// TIA Portal project "Tank_Level_FactoryIO" (V15.1)

(* hardware
DEVICE "S7-1200 station_1"  S7-1200 Station
   slot 0: "Rack_0"  S7-1200 Rack  Rack  V1.0
   slot 1: "PLC_1"  CPU 1214C DC/DC/DC  6ES7 214-1AG40-0XB0  V4.2
DEVICE "HMI_1"  TP1500 Comfort PRO
   slot 0: "HMI_1"  TP1500 Comfort PRO  6AV2 124-0QC24-1AX0  15.1.0.0
   slot 1: "HMI_RT_1"  TP1500 Comfort PRO  6AV2 124-0QC24-1AX0  15.1.0.0
   slot 5: "HMI_1.IE_CP_1"  PROFINET Interface  15.0.1.0
      slot 1: "PROFINET Interface_1"  PROFINET Interface
         slot 1: "Port_1"  Port
         slot 2: "Port_2"  Port
   slot 6: "HMI_1.IE_CP_2"  PROFINET Interface  15.0.1.0
      slot 1: "PROFINET Interface_GBit"  PROFINET Interface
         slot 1: "Port_1"  Port
   slot 7: "HMI_1.MPI/DP_CP_1"  MPI/DP Interface  15.0.1.0
*)

// ===== PLC "PLC_1"  CPU 1214C DC/DC/DC =====

VAR_GLOBAL   // PLC tag table "Default tag table"
   "Raw_Sensor_Sim" AT %MW10 : Int;
   "Level_Normalized" AT %MD20 : Real;
   "Level_CM" AT %MD24 : Real;
   "Fill_Valve" AT %QW30 : Int;
   "Pump_Cmd" AT %Q0.0 : Bool;
   "I_Start" AT %I0.0 : Bool;
   "I_Stop" AT %I0.1 : Bool;
   "System_Active" AT %M0.0 : Bool;
   "Discharge_Valve" AT %Q0.1 : Bool;
   "Sim_Tick" AT %M50.0 : Bool;
   "Level_Input_Raw" AT %IW30 : Int;
   "Discharge_Valve_Analog" AT %QW32 : Int;
   "HMI_Start" AT %M10.0 : Bool;
   "HMI_Stop" AT %M12.0 : Bool;
END_VAR

FUNCTION "Signal Conversion" : Void   // FC1, LAD
{ S7_Optimized_Access := 'TRUE' }
VERSION : 0.1
BEGIN

REGION Network 1: Signal Conversion
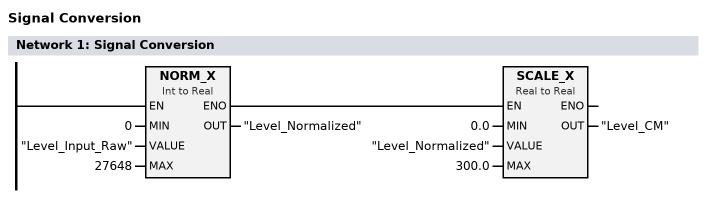
   RUNG wire#powerrail
      { S7_Templates := "[SrcType := Int, DestType := Real]" } Normalize(min := 0, value := "Level_Input_Raw", max := 27648, out => "Level_Normalized")
      { S7_Templates := "[SrcType := Real, DestType := Real]" } Scale(min := 0.0, value := "Level_Normalized", max := 300.0, out => "Level_CM")
   END_RUNG
   // the same network as SCL:
   "Level_Normalized" := NORM_X(MIN := 0, VALUE := "Level_Input_Raw", MAX := 27648);
   "Level_CM" := SCALE_X(MIN := 0.0, VALUE := "Level_Normalized", MAX := 300.0);
END_REGION
END_FUNCTION

FUNCTION "Pump Control" : Void   // FC2, LAD
{ S7_Optimized_Access := 'TRUE' }
VERSION : 0.1
BEGIN

REGION Network 1
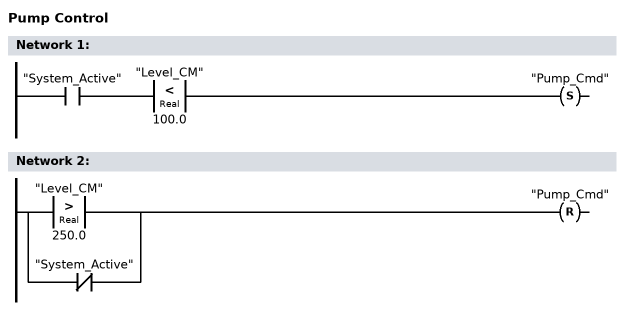
   RUNG wire#powerrail
      Contact( "System_Active" )
      { S7_Templates := "SrcType := Real" } LT_Contact(in1 := "Level_CM", in2 := 100.0)
      S_Coil( "Pump_Cmd" )
   END_RUNG
   // the same network as SCL:
   IF "System_Active" AND ("Level_CM" < 100.0) THEN "Pump_Cmd" := TRUE; END_IF;
END_REGION

REGION Network 2
   RUNG wire#powerrail
      { S7_Templates := "SrcType := Real" } GT_Contact(in1 := "Level_CM", in2 := 250.0)
      wire#w1
      R_Coil( "Pump_Cmd" )
   END_RUNG
   RUNG wire#powerrail
      I_Contact( "System_Active" )
   END_RUNG wire#w1
   // the same network as SCL:
   IF ("Level_CM" > 250.0) OR NOT "System_Active" THEN "Pump_Cmd" := FALSE; END_IF;
END_REGION
END_FUNCTION

FUNCTION "Discharge Valve" : Void   // FC3, LAD
{ S7_Optimized_Access := 'TRUE' }
VERSION : 0.1
BEGIN

REGION Network 1
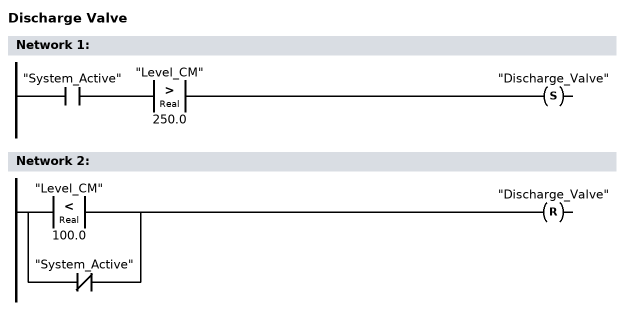
   RUNG wire#powerrail
      Contact( "System_Active" )
      { S7_Templates := "SrcType := Real" } GT_Contact(in1 := "Level_CM", in2 := 250.0)
      S_Coil( "Discharge_Valve" )
   END_RUNG
   // the same network as SCL:
   IF "System_Active" AND ("Level_CM" > 250.0) THEN "Discharge_Valve" := TRUE; END_IF;
END_REGION

REGION Network 2
   RUNG wire#powerrail
      { S7_Templates := "SrcType := Real" } LT_Contact(in1 := "Level_CM", in2 := 100.0)
      wire#w1
      R_Coil( "Discharge_Valve" )
   END_RUNG
   RUNG wire#powerrail
      I_Contact( "System_Active" )
   END_RUNG wire#w1
   // the same network as SCL:
   IF ("Level_CM" < 100.0) OR NOT "System_Active" THEN "Discharge_Valve" := FALSE; END_IF;
END_REGION
END_FUNCTION

FUNCTION "MHJ-PLC-Lab-Function-S71200" : Void   // FC9000, SCL
{ S7_Optimized_Access := 'TRUE' }
VERSION : 0.1
   VAR_TEMP
      rdTimeReturn : Int;
      outputTime : DTL;
      SyncVal : Byte;
      forVal : Int;
      forVal_2 : Int;
      Value : Byte;
   END_VAR
   VAR CONSTANT
      CompVal : Byte := 16#34;
      Value_01 : Byte := 16#11;
      Value_01_DW : DWord := 16#A165_D992;
      Value_02_DW : DWord := 16#58BE_4401;
   END_VAR
BEGIN

   #Value:=PEEK(area := 16#82,
        dbNumber := 0,
        byteOffset := 511);
   #Value := #Value + 1;

   POKE(area := 16#82,
        dbNumber := 0,
        byteOffset := 511,
        value := #Value);

   POKE(area:=16#81,
        dbNumber:=0,
        byteOffset:=1016,
        value:=#Value_01_DW);
   POKE(area := 16#81,
        dbNumber := 0,
        byteOffset := 1020,
        value := #Value_02_DW);

   POKE(area := 16#81,
        dbNumber := 0,
        byteOffset := 511,
        value := B#16#00);

   FOR #forVal := 0 TO 120 DO
       FOR #forVal_2:=0 TO 10 DO
           #rdTimeReturn:=RD_SYS_T(#outputTime);
           #rdTimeReturn := WR_SYS_T(#outputTime);
           #rdTimeReturn := RD_SYS_T(#outputTime);
           #rdTimeReturn := WR_SYS_T(#outputTime);
       END_FOR;
       #SyncVal:= PEEK(area := 16#81,
                      dbNumber := 0,
                      byteOffset := 511);
       IF #SyncVal = #CompVal THEN
          GOTO M_1;
       END_IF;
   END_FOR;
   RETURN;

   M_1:
   POKE(area := 16#81,
        dbNumber := 0,
        byteOffset := 511,
        value := B#16#0);
END_FUNCTION

ORGANIZATION_BLOCK "Main"   // OB1, LAD, ProgramCycle
TITLE = "Main Program Sweep (Cycle)"
{ S7_Optimized_Access := 'TRUE' }
VERSION : 0.1
   VAR_INPUT
      Initial_Call : Bool;   // Initial call of this OB
      Remanence : Bool;   // =True, if remanent data are available
   END_VAR
BEGIN

REGION Network 1: Factory I/O Setup Template
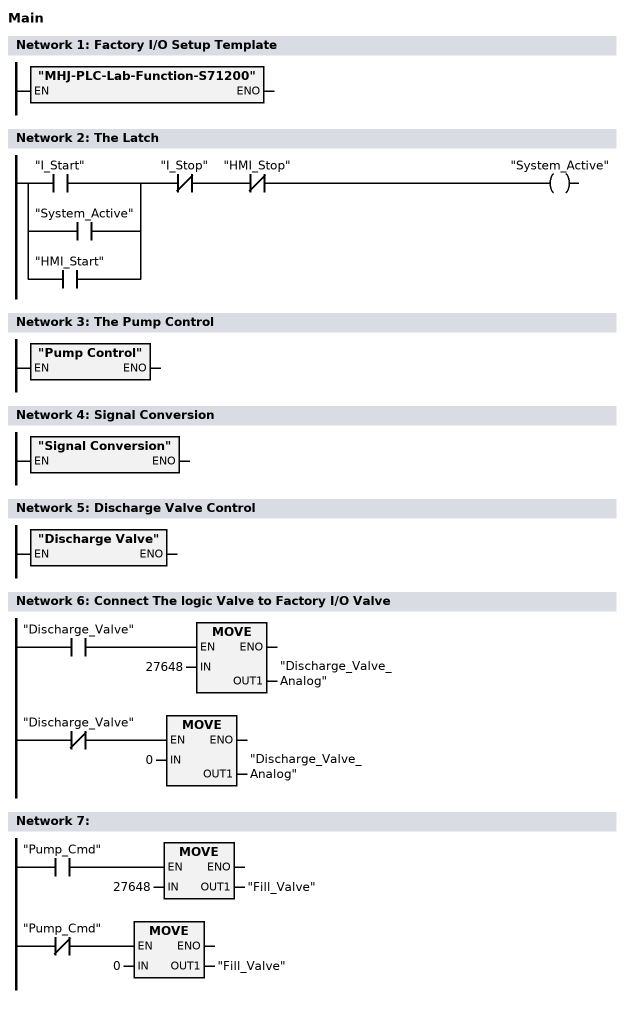
   RUNG wire#powerrail
      "MHJ-PLC-Lab-Function-S71200"()
   END_RUNG
   // the same network as SCL:
   "MHJ-PLC-Lab-Function-S71200"();
END_REGION

REGION Network 2: The Latch
   RUNG wire#powerrail
      Contact( "I_Start" )
      wire#w1
      I_Contact( "I_Stop" )
      I_Contact( "HMI_Stop" )
      Coil( "System_Active" )
   END_RUNG
   RUNG wire#powerrail
      Contact( "System_Active" )
   END_RUNG wire#w1
   RUNG wire#powerrail
      Contact( "HMI_Start" )
   END_RUNG wire#w1
   // the same network as SCL:
   "System_Active" := ("I_Start" OR "System_Active" OR "HMI_Start") AND NOT "I_Stop" AND NOT "HMI_Stop";
END_REGION

REGION Network 3: The Pump Control
   RUNG wire#powerrail
      "Pump Control"()
   END_RUNG
   // the same network as SCL:
   "Pump Control"();
END_REGION

REGION Network 4: Signal Conversion
   RUNG wire#powerrail
      "Signal Conversion"()
   END_RUNG
   // the same network as SCL:
   "Signal Conversion"();
END_REGION

REGION Network 5: Discharge Valve Control
   RUNG wire#powerrail
      "Discharge Valve"()
   END_RUNG
   // the same network as SCL:
   "Discharge Valve"();
END_REGION

REGION Network 6: Connect The logic Valve to Factory I/O Valve
   RUNG wire#powerrail
      Contact( "Discharge_Valve" )
      Move(in := 27648, out1 => "Discharge_Valve_Analog")
   END_RUNG
   RUNG wire#powerrail
      I_Contact( "Discharge_Valve" )
      Move(in := 0, out1 => "Discharge_Valve_Analog")
   END_RUNG
   // the same network as SCL:
   IF "Discharge_Valve" THEN "Discharge_Valve_Analog" := 27648; END_IF;
   IF NOT "Discharge_Valve" THEN "Discharge_Valve_Analog" := 0; END_IF;
END_REGION

REGION Network 7
   RUNG wire#powerrail
      Contact( "Pump_Cmd" )
      Move(in := 27648, out1 => "Fill_Valve")
   END_RUNG
   RUNG wire#powerrail
      I_Contact( "Pump_Cmd" )
      Move(in := 0, out1 => "Fill_Valve")
   END_RUNG
   // the same network as SCL:
   IF "Pump_Cmd" THEN "Fill_Valve" := 27648; END_IF;
   IF NOT "Pump_Cmd" THEN "Fill_Valve" := 0; END_IF;
END_REGION
END_ORGANIZATION_BLOCK

(* ===== HMI "HMI_RT_1" =====
system functions are stored by id; their names below are inferred from use
connection "HMI_Connection_1": ETHERNET, S7_1200_OMS

HMI tags "Default tag table"
   "Tag_ScreenNumber" : UInt, internal
   "Raw_Sensor_Sim" : Int = PLC Raw_Sensor_Sim AT %MW10, 1 s
   "Level_CM" : Real = PLC Level_CM AT %MD24, 1 s
   "Pump_Cmd" : Bool = PLC Pump_Cmd AT %Q0.0, 1 s
   "Discharge_Valve" : Bool = PLC Discharge_Valve AT %Q0.1, 1 s
   "Fill_Valve" : Int = PLC Fill_Valve AT %QW30, 1 s
   "HMI_Start" : Bool = PLC HMI_Start AT %M10.0, 1 s
   "HMI_Stop" : Bool = PLC HMI_Stop AT %M12.0, 1 s
   "Level_Input_Raw" : Int = PLC Level_Input_Raw AT %IW30, 1 s

screen "Root screen" 1366x708, template "Template_1"
   on GenerateScreen: SetTag("Tag_ScreenNumber", 1)
   Bar "Bar_1" at 1126,327 size 80x230; MinimumValue 0; MaximumValue 300
      ProcessValue <- "Level_CM"
   Circle "Circle_1" at 1247,100 size 48x48
      Appearance <- "Pump_Cmd"
   TextField "Text field_1" at 472,9 size 322x58; Text 'Tank Supervisor'
   GraphicView "Graphic view_1" at 1011,67 size 211x98; Picture "Graphic_1"
   GraphicView "Graphic view_2" at 1036,188 size 190x103; Picture "Graphic_2"
   Circle "Circle_2" at 1247,222 size 48x48
      Appearance <- "Discharge_Valve"
   TextField "Text field_2" at 985,569 size 334x58; Text 'Tank Level in CM'
   TextField "Text field_3" at 272,562 size 275x58; Text 'Sensor Reads'
   Group "Group" at 862,96 size 115x52
   Group "Group_1" at 856,213 size 154x63
   Button "Button_1" at 100,325 size 132x63; TextOff 'START'
      on Press: function_b14e0dd5("HMI_Start", 0)
   Button "Button_2" at 101,446 size 132x63; TextOff 'STOP'
      on Press: function_b14e0dd5("HMI_Stop", 0)
   Bar "Bar_2" at 372,316 size 80x230; MinimumValue 0; MaximumValue 27648
      ProcessValue <- "Level_Input_Raw"
   TextField "Text field_4" at 888,107 size 58x25; Text 'Pump'
   TextField "Text field_5" at 885,222 size 106x46; Text 'Discharge Valve'

Template "Template_1" 1366x708
   Button "Exit" at 1286,647 size 78x59; TextOff 'Exit'; PictureOff "ExitRuntime_TP1500_Comfort_PRO_TR"; PictureOn "ExitRuntime_TP1500_Comfort_PRO_TR"
      on Release: StopRuntime(0)
   Button "Template_Button" at 1205,647 size 78x59; TextOff 'Text'
   Button "Template_Button_1" at 1125,647 size 78x59; TextOff 'Text'
   Button "Template_Button_2" at 1045,647 size 78x59; TextOff 'Text'
   Button "Template_Button_3" at 965,647 size 78x59; TextOff 'Text'
   Button "Template_Button_4" at 884,647 size 78x59; TextOff 'Text'
   Button "Template_Button_5" at 804,647 size 78x59; TextOff 'Text'
   Button "Template_Button_6" at 724,647 size 78x59; TextOff 'Text'
   Button "Template_Button_7" at 643,647 size 78x59; TextOff 'Text'
   Button "Template_Button_8" at 563,647 size 78x59; TextOff 'Text'
   Button "Template_Button_9" at 483,647 size 78x59; TextOff 'Text'
   Button "Template_Button_10" at 402,647 size 78x59; TextOff 'Text'
   Button "Template_Button_11" at 322,647 size 78x59; TextOff 'Text'
   Button "Template_Button_12" at 242,647 size 78x59; TextOff 'Text'
   Button "Template_Button_13" at 162,647 size 78x59; TextOff 'Text'
   Button "Template_Button_14" at 81,647 size 78x59; TextOff 'Text'
   Button "Start screen" at 1,647 size 78x59; TextOff 'Start screen'; PictureOff "NavigateHome_TP1500_Comfort_PRO_TR"; PictureOn "NavigateHome_TP1500_Comfort_PRO_TR"
      on Release: ActivateScreen("Root screen", 0)
*)